(* Logix 5000 project; controller _GigaDiscovery vendor 1 type 14 code 244 rev 35.11; software revision 35.03; part 16 of 23 *)
(* tags used below, declared in another part *)
   E_Stop2_Test_Request : BOOL;
   E_Stop_Test_Request : BOOL;
   HMI_Pb_Platform_Open : BOOL;   // HMI Platform Open Command
   HMI_Platform_Close : BOOL;   // HMI Platform Close Command
   I_Compressor_Min_Pressure : BOOL;   // Line Pressure Switch - Minimum Pressure -S21504B
   I_Compressor_Work_Pressure : BOOL;   // Line Pressure Switch - Working Pressure -S21502B
   I_EStop_Pb_OCC1 : UDT_DCI_STOP_TEST;   // +OCC E-stop -S30301F
   I_EStop_Pb_OCC2 : UDT_DCI_STOP_TEST;   // +OCC2 E-Stop -S28502F
   I_HMI_Login_Enable : BOOL;   // Primary console Key selector Display Login -S30309F
   I_MCC_Temperature_OK : BOOL;   // MCC temeprature OK -S75003C
   I_OCC1_EntGate_PB : BOOL;   // OCC1 Entrance Gate Open/Close -S30701F
   I_OCC1_ExitGate_PB : BOOL;   // OCC1 ExitGate Open/Close -S30707F
   I_OCC1_Stop_Cycle_PB : BOOL;   // Stop Cycle -S30308F
   I_OCC2_ACONFIRM : BOOL;   // OCC2 Allow Main CONFIRM -S28602F
   I_OCC2_Disable : UDT_DCM;   // OCC 2 CONTROL DISABLE Page 310
   I_OCC2_RESTRAINTS_RELEASE : Sel_3_Pos_2_Input;   // -S28507F RESTRAINTS RELEASE UNLOCK -RUN- LOCK
   I_OCC2_Stop_Cycle_PB : BOOL;   // Stop Cycle -S28606F
   I_OCC_Aut_Man_Selector_Motion : UDT_DCM;   // S30801F
   I_OCC_Emergency_Brake : BOOL;   // I OCC Emergency Brake -S31207D
   I_OCC_LockOut_Motion : UDT_DCM;   // OCC -Lockout Motion -Q31203E
   I_OCC_Memory_Footpedal : BOOL;
   I_OCC_Operator_Enable_Key : BOOL;   // OCC Console Enabled -S30305F
   I_OCC_Temperature_OK : BOOL;   // OCC temperature OK -S31003E
   I_Operator_Footpedal : BOOL;   // Operator Footpedal -S30901F
   I_RESTRAINTS_MainValve_Cosed : BOOL;   // Main Valve Close Limit Switch -B40508I
   I_RESTRAINTS_PressureswitchCompressor : BOOL;   // RESTRAINTS Main Valve Pressure Switch -S40602J
   I_RESTRAINTS_Selector : Sel_3_Pos_2_Input;   // RESTRAINTS Selctor -S30505F Left = Open Right = Close Center = Nothing
   I_Start_PB : Start_AOI;   // Primary console Strat Push botton Right and Left -S30401F -S30403F
   MODE : BOOL;   // MODE 0 = AUTO 1 = MANUAL -S30801F
   No_Sfty : Std_to_Sfty;
   ONP : DINT;   // Optional Not Present
   Pb_Platform_Stop : BOOL;   // Platform Stop Command -S30608F
   Power_On_Delay : BOOL;
   Reset_Pulse : BOOL;
   RESTRAINTS_Rack : LapBar_Racks[41];
   RESTRAINTS_Sector : LapBars_Sector[9];
   Start_Stop_Cycle : Sequencer;
   ToBe_Define_Sfty : DINT[10];

PROGRAM S_Input   (* main routine Main, safety *)
VAR
   E_Stop_Secondary_Released : BOOL := 1;
   Home_Timer : TIMER := (PRE := 10000, ACC := 10000, EN := 1, DN := 1);
   Os : DINT := 14;
   Reset_Start_AOI : BOOL;   // Start AOI Instruction Reset
   Reset_Status : TIMER := (PRE := 1500, ACC := 1520);
   timer : TIMER[10] := ([0].PRE := 30000, [0].ACC := 30000, [0].EN := 1, [0].DN := 1, [1].PRE := 8000, [1].ACC := 8000, [1].EN := 1, [1].DN := 1, [2].PRE := 3000, [2].EN := 1, [2].DN := 1, [3].PRE := 4000, [4].PRE := 2000, [5].PRE := 5000, [6].PRE := 500, [7].PRE := 500, [8].PRE := 1600);
   Timer2 : TIMER := (PRE := 5000, ACC := 5000, EN := 1, DN := 1);
END_VAR

ROUTINE _01_OCC   (* ladder *)
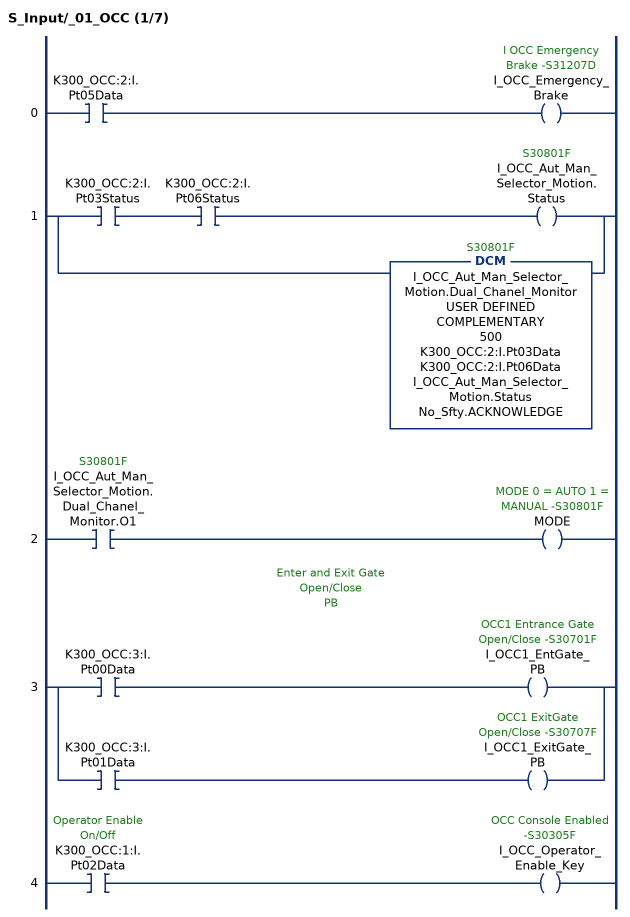
   0: XIC(K300_OCC:2:I.Pt05Data)OTE(I_OCC_Emergency_Brake);
   1: [XIC(K300_OCC:2:I.Pt03Status) XIC(K300_OCC:2:I.Pt06Status) OTE(I_OCC_Aut_Man_Selector_Motion.Status) ,DCM(I_OCC_Aut_Man_Selector_Motion.Dual_Chanel_Monitor,USER DEFINED,COMPLEMENTARY,500,K300_OCC:2:I.Pt03Data,K300_OCC:2:I.Pt06Data,I_OCC_Aut_Man_Selector_Motion.Status,No_Sfty.ACKNOWLEDGE) ];
   2: XIC(I_OCC_Aut_Man_Selector_Motion.Dual_Chanel_Monitor.O1)OTE(MODE);
   // Enter and Exit Gate
   // Open/Close
   // PB
   3: [XIC(K300_OCC:3:I.Pt00Data) OTE(I_OCC1_EntGate_PB) ,XIC(K300_OCC:3:I.Pt01Data) OTE(I_OCC1_ExitGate_PB) ];
   4: XIC(K300_OCC:1:I.Pt02Data)OTE(I_OCC_Operator_Enable_Key);
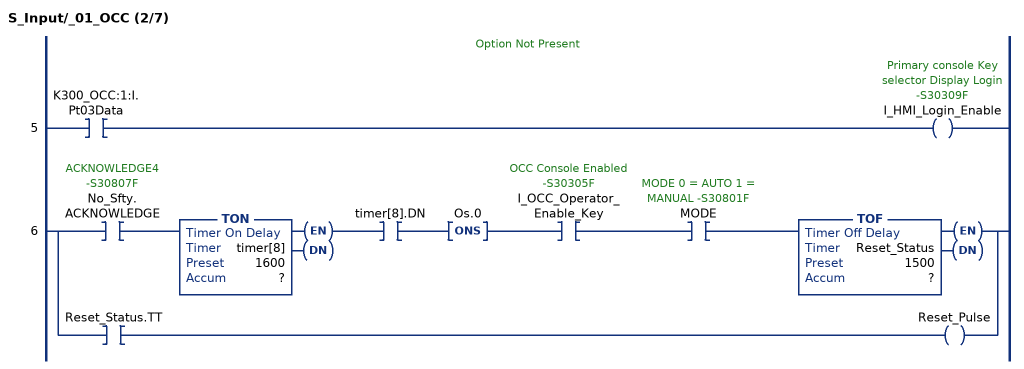
   // Option Not Present
   5: XIC(K300_OCC:1:I.Pt03Data)OTE(I_HMI_Login_Enable);
   6: [XIC(No_Sfty.ACKNOWLEDGE) TON(timer[8],?,?) XIC(timer[8].DN) ONS(Os.0) XIC(I_OCC_Operator_Enable_Key) XIC(MODE) TOF(Reset_Status,?,?) ,XIC(Reset_Status.TT) OTE(Reset_Pulse) ];
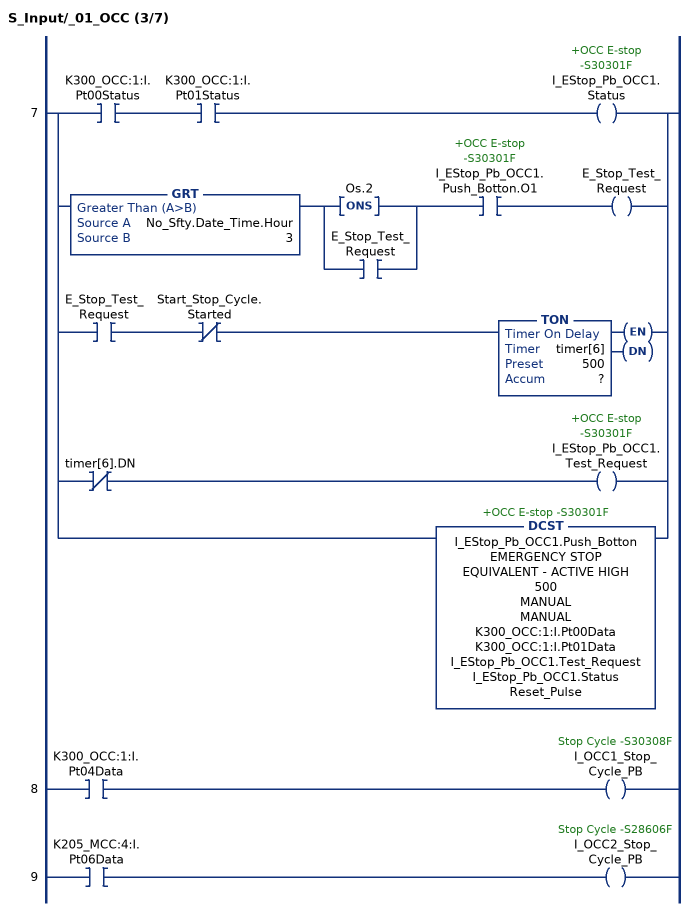
   7: [XIC(K300_OCC:1:I.Pt00Status) XIC(K300_OCC:1:I.Pt01Status) OTE(I_EStop_Pb_OCC1.Status) ,GRT(No_Sfty.Date_Time.Hour,3) [ONS(Os.2) ,XIC(E_Stop_Test_Request) ] XIC(I_EStop_Pb_OCC1.Push_Botton.O1) OTE(E_Stop_Test_Request) ,XIC(E_Stop_Test_Request) XIO(Start_Stop_Cycle.Started) TON(timer[6],?,?) ,XIO(timer[6].DN) OTE(I_EStop_Pb_OCC1.Test_Request) ,DCST(I_EStop_Pb_OCC1.Push_Botton,EMERGENCY STOP,EQUIVALENT - ACTIVE HIGH,500,MANUAL,MANUAL,K300_OCC:1:I.Pt00Data,K300_OCC:1:I.Pt01Data,I_EStop_Pb_OCC1.Test_Request,I_EStop_Pb_OCC1.Status,Reset_Pulse) ];
   8: XIC(K300_OCC:1:I.Pt04Data)OTE(I_OCC1_Stop_Cycle_PB);
   9: XIC(K205_MCC:4:I.Pt06Data)OTE(I_OCC2_Stop_Cycle_PB);
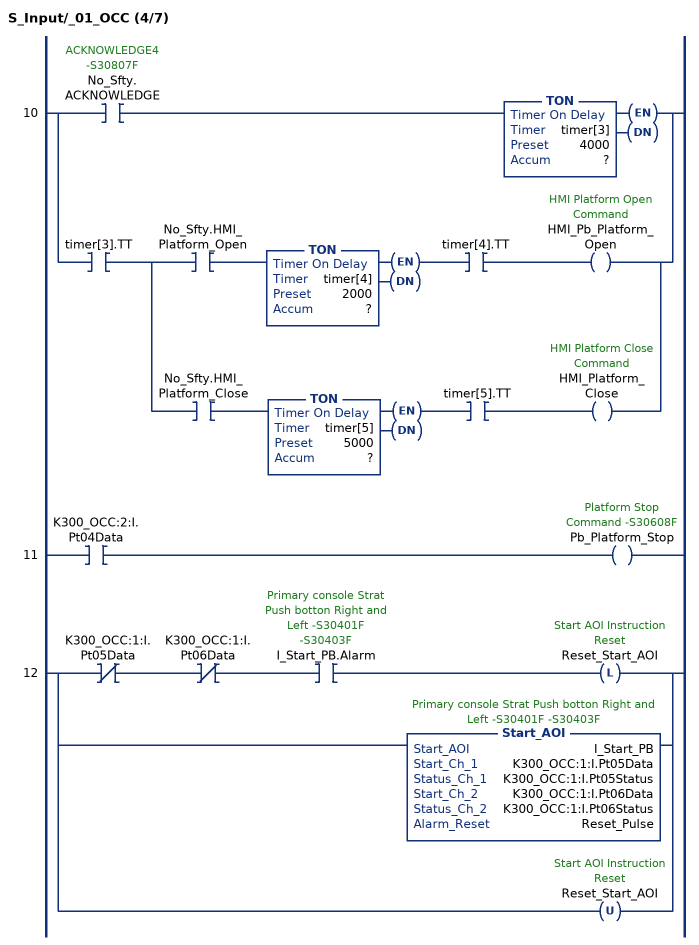
   10: [XIC(No_Sfty.ACKNOWLEDGE) TON(timer[3],?,?) ,XIC(timer[3].TT) [XIC(No_Sfty.HMI_Platform_Open) TON(timer[4],?,?) XIC(timer[4].TT) OTE(HMI_Pb_Platform_Open) ,XIC(No_Sfty.HMI_Platform_Close) TON(timer[5],?,?) XIC(timer[5].TT) OTE(HMI_Platform_Close) ] ];
   11: XIC(K300_OCC:2:I.Pt04Data)OTE(Pb_Platform_Stop);
   12: [XIO(K300_OCC:1:I.Pt05Data) XIO(K300_OCC:1:I.Pt06Data) XIC(I_Start_PB.Alarm) OTL(Reset_Start_AOI) ,Start_AOI(I_Start_PB,K300_OCC:1:I.Pt05Data,K300_OCC:1:I.Pt05Status,K300_OCC:1:I.Pt06Data,K300_OCC:1:I.Pt06Status,Reset_Pulse) ,OTU(Reset_Start_AOI) ];
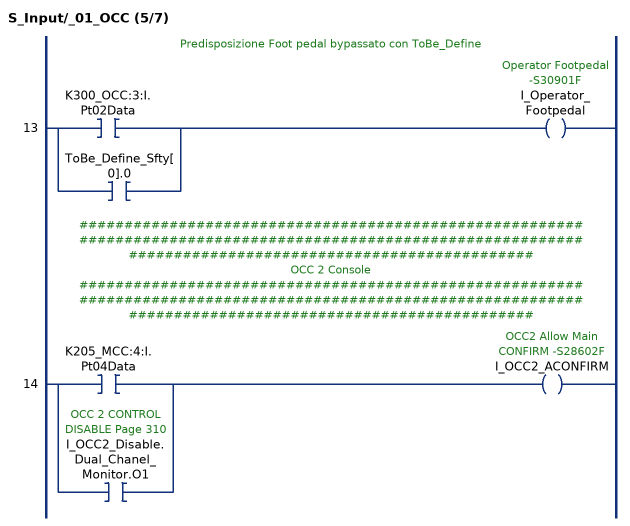
   // Predisposizione Foot pedal bypassato con ToBe_Define
   13: [XIC(K300_OCC:3:I.Pt02Data) ,XIC(ToBe_Define_Sfty[0].0) ]OTE(I_Operator_Footpedal);
   // #############################################################################################################################################################
   // OCC 2 Console
   // #############################################################################################################################################################
   14: [XIC(K205_MCC:4:I.Pt04Data) ,XIC(I_OCC2_Disable.Dual_Chanel_Monitor.O1) ]OTE(I_OCC2_ACONFIRM);
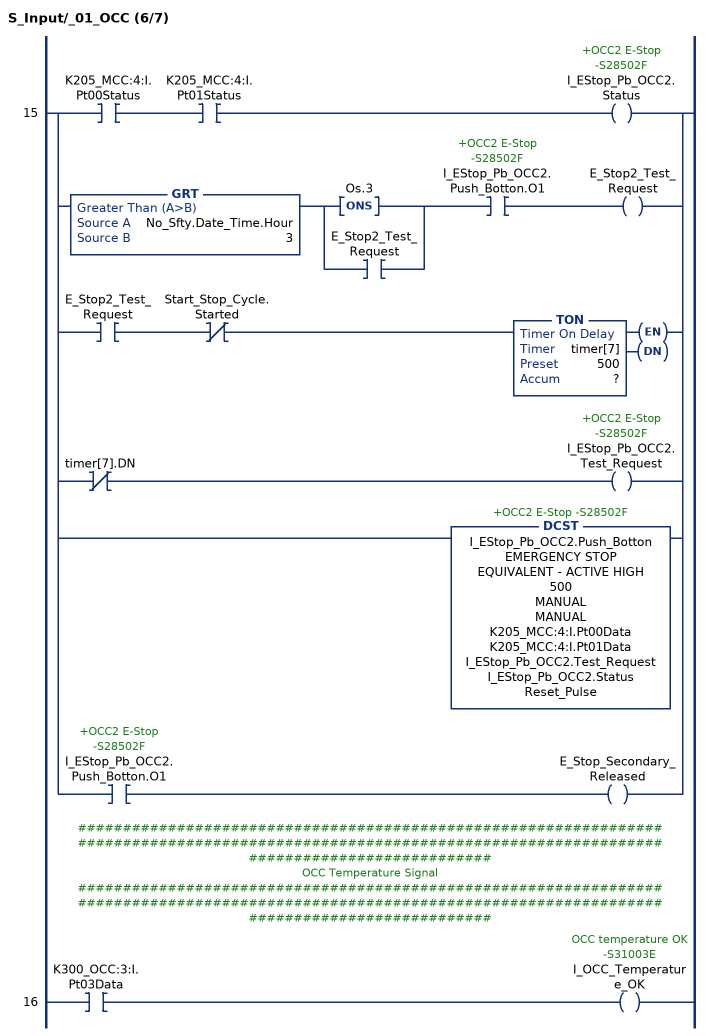
   15: [XIC(K205_MCC:4:I.Pt00Status) XIC(K205_MCC:4:I.Pt01Status) OTE(I_EStop_Pb_OCC2.Status) ,GRT(No_Sfty.Date_Time.Hour,3) [ONS(Os.3) ,XIC(E_Stop2_Test_Request) ] XIC(I_EStop_Pb_OCC2.Push_Botton.O1) OTE(E_Stop2_Test_Request) ,XIC(E_Stop2_Test_Request) XIO(Start_Stop_Cycle.Started) TON(timer[7],?,?) ,XIO(timer[7].DN) OTE(I_EStop_Pb_OCC2.Test_Request) ,DCST(I_EStop_Pb_OCC2.Push_Botton,EMERGENCY STOP,EQUIVALENT - ACTIVE HIGH,500,MANUAL,MANUAL,K205_MCC:4:I.Pt00Data,K205_MCC:4:I.Pt01Data,I_EStop_Pb_OCC2.Test_Request,I_EStop_Pb_OCC2.Status,Reset_Pulse) ,XIC(I_EStop_Pb_OCC2.Push_Botton.O1) OTE(E_Stop_Secondary_Released) ];
   // #############################################################################################################################################################
   // OCC Temperature Signal
   // #############################################################################################################################################################
   16: XIC(K300_OCC:3:I.Pt03Data)OTE(I_OCC_Temperature_OK);
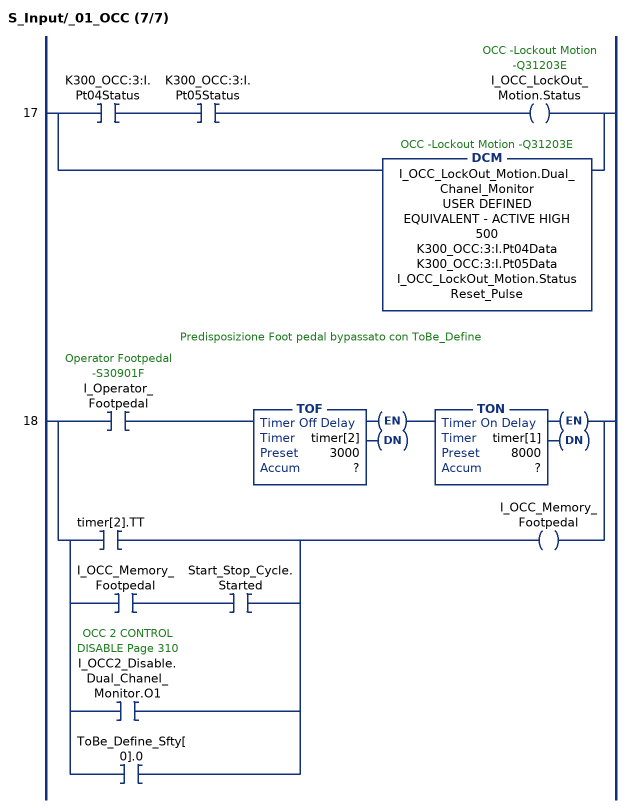
   17: [XIC(K300_OCC:3:I.Pt04Status) XIC(K300_OCC:3:I.Pt05Status) OTE(I_OCC_LockOut_Motion.Status) ,DCM(I_OCC_LockOut_Motion.Dual_Chanel_Monitor,USER DEFINED,EQUIVALENT - ACTIVE HIGH,500,K300_OCC:3:I.Pt04Data,K300_OCC:3:I.Pt05Data,I_OCC_LockOut_Motion.Status,Reset_Pulse) ];
   // Predisposizione Foot pedal bypassato con ToBe_Define
   18: [XIC(I_Operator_Footpedal) TOF(timer[2],?,?) TON(timer[1],?,?) ,[XIC(timer[2].TT) ,XIC(I_OCC_Memory_Footpedal) XIC(Start_Stop_Cycle.Started) ,XIC(I_OCC2_Disable.Dual_Chanel_Monitor.O1) ,XIC(ToBe_Define_Sfty[0].0) ] OTE(I_OCC_Memory_Footpedal) ];
END_ROUTINE

ROUTINE _02_MCC   (* ladder *)
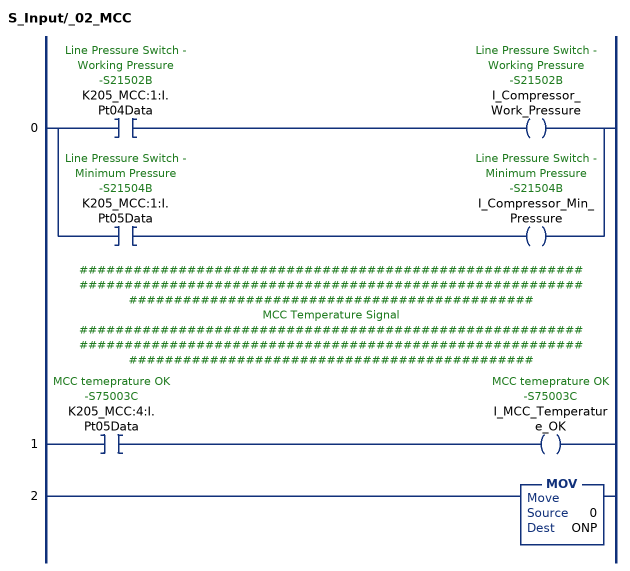
   0: [XIC(K205_MCC:1:I.Pt04Data) OTE(I_Compressor_Work_Pressure) ,XIC(K205_MCC:1:I.Pt05Data) OTE(I_Compressor_Min_Pressure) ];
   // #############################################################################################################################################################
   // MCC Temperature Signal
   // #############################################################################################################################################################
   1: XIC(K205_MCC:4:I.Pt05Data)OTE(I_MCC_Temperature_OK);
   2: MOV(0,ONP);
END_ROUTINE

ROUTINE _03_RESTRAINT_RELEASE   (* ladder *)
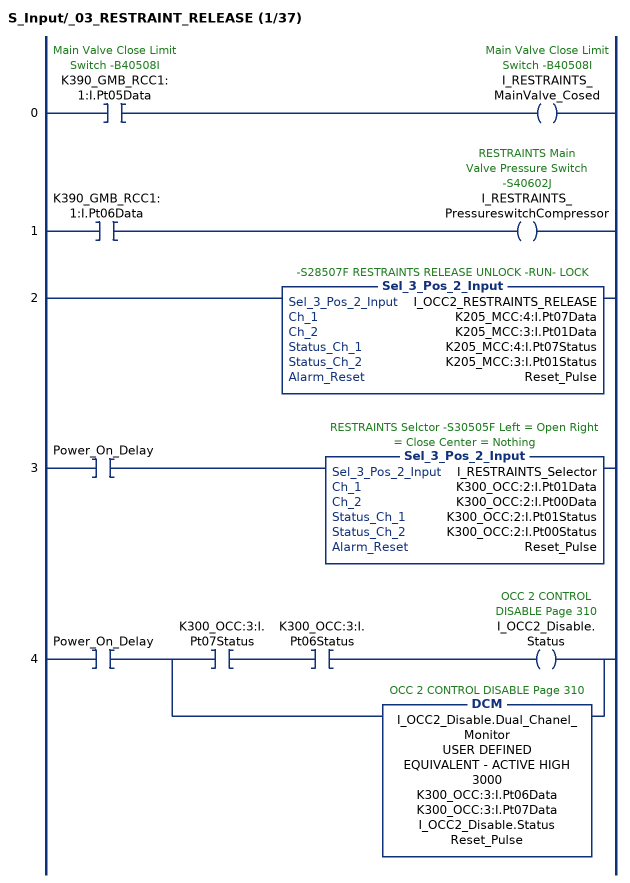
   0: XIC(K390_GMB_RCC1:1:I.Pt05Data)OTE(I_RESTRAINTS_MainValve_Cosed);
   1: XIC(K390_GMB_RCC1:1:I.Pt06Data)OTE(I_RESTRAINTS_PressureswitchCompressor);
   2: Sel_3_Pos_2_Input(I_OCC2_RESTRAINTS_RELEASE,K205_MCC:4:I.Pt07Data,K205_MCC:3:I.Pt01Data,K205_MCC:4:I.Pt07Status,K205_MCC:3:I.Pt01Status,Reset_Pulse);
   3: XIC(Power_On_Delay)Sel_3_Pos_2_Input(I_RESTRAINTS_Selector,K300_OCC:2:I.Pt01Data,K300_OCC:2:I.Pt00Data,K300_OCC:2:I.Pt01Status,K300_OCC:2:I.Pt00Status,Reset_Pulse);
   4: XIC(Power_On_Delay)[XIC(K300_OCC:3:I.Pt07Status) XIC(K300_OCC:3:I.Pt06Status) OTE(I_OCC2_Disable.Status) ,DCM(I_OCC2_Disable.Dual_Chanel_Monitor,USER DEFINED,EQUIVALENT - ACTIVE HIGH,3000,K300_OCC:3:I.Pt06Data,K300_OCC:3:I.Pt07Data,I_OCC2_Disable.Status,Reset_Pulse) ];
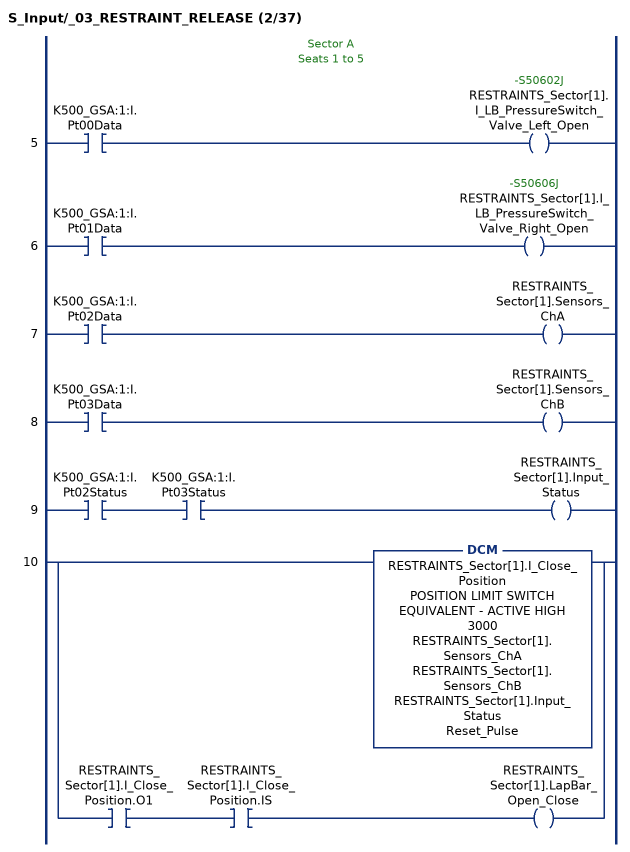
   // Sector A
   // Seats 1 to 5
   5: XIC(K500_GSA:1:I.Pt00Data)OTE(RESTRAINTS_Sector[1].I_LB_PressureSwitch_Valve_Left_Open);
   6: XIC(K500_GSA:1:I.Pt01Data)OTE(RESTRAINTS_Sector[1].I_LB_PressureSwitch_Valve_Right_Open);
   7: XIC(K500_GSA:1:I.Pt02Data)OTE(RESTRAINTS_Sector[1].Sensors_ChA);
   8: XIC(K500_GSA:1:I.Pt03Data)OTE(RESTRAINTS_Sector[1].Sensors_ChB);
   9: XIC(K500_GSA:1:I.Pt02Status)XIC(K500_GSA:1:I.Pt03Status)OTE(RESTRAINTS_Sector[1].Input_Status);
   10: [DCM(RESTRAINTS_Sector[1].I_Close_Position,POSITION LIMIT SWITCH,EQUIVALENT - ACTIVE HIGH,3000,RESTRAINTS_Sector[1].Sensors_ChA,RESTRAINTS_Sector[1].Sensors_ChB,RESTRAINTS_Sector[1].Input_Status,Reset_Pulse) ,XIC(RESTRAINTS_Sector[1].I_Close_Position.O1) XIC(RESTRAINTS_Sector[1].I_Close_Position.IS) OTE(RESTRAINTS_Sector[1].LapBar_Open_Close) ];
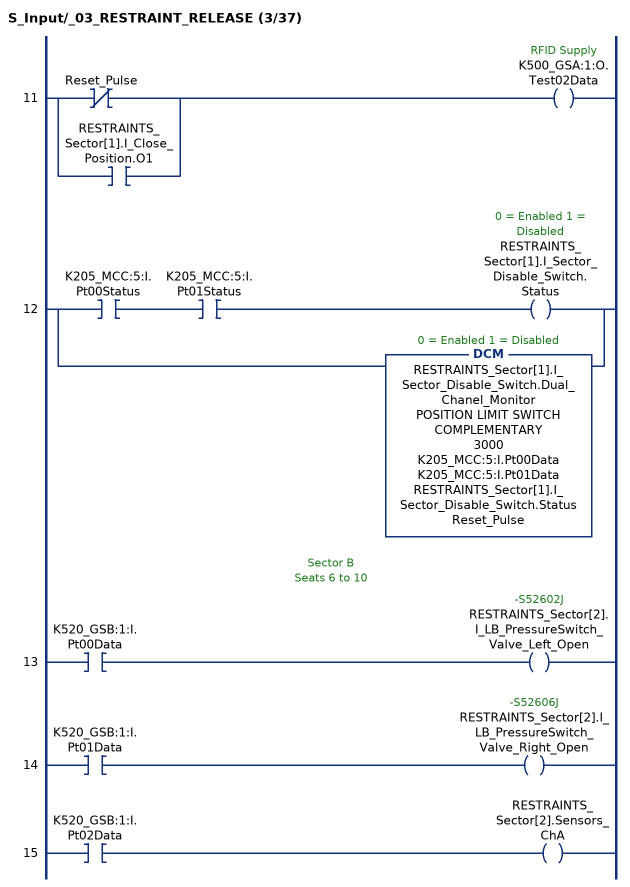
   11: [XIO(Reset_Pulse) ,XIC(RESTRAINTS_Sector[1].I_Close_Position.O1) ]OTE(K500_GSA:1:O.Test02Data);
   12: [XIC(K205_MCC:5:I.Pt00Status) XIC(K205_MCC:5:I.Pt01Status) OTE(RESTRAINTS_Sector[1].I_Sector_Disable_Switch.Status) ,DCM(RESTRAINTS_Sector[1].I_Sector_Disable_Switch.Dual_Chanel_Monitor,POSITION LIMIT SWITCH,COMPLEMENTARY,3000,K205_MCC:5:I.Pt00Data,K205_MCC:5:I.Pt01Data,RESTRAINTS_Sector[1].I_Sector_Disable_Switch.Status,Reset_Pulse) ];
   // Sector B
   // Seats 6 to 10
   13: XIC(K520_GSB:1:I.Pt00Data)OTE(RESTRAINTS_Sector[2].I_LB_PressureSwitch_Valve_Left_Open);
   14: XIC(K520_GSB:1:I.Pt01Data)OTE(RESTRAINTS_Sector[2].I_LB_PressureSwitch_Valve_Right_Open);
   15: XIC(K520_GSB:1:I.Pt02Data)OTE(RESTRAINTS_Sector[2].Sensors_ChA);
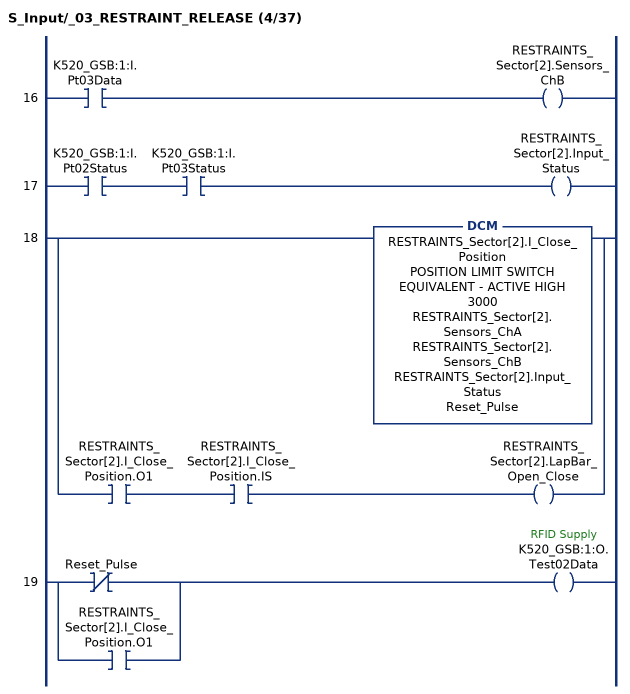
   16: XIC(K520_GSB:1:I.Pt03Data)OTE(RESTRAINTS_Sector[2].Sensors_ChB);
   17: XIC(K520_GSB:1:I.Pt02Status)XIC(K520_GSB:1:I.Pt03Status)OTE(RESTRAINTS_Sector[2].Input_Status);
   18: [DCM(RESTRAINTS_Sector[2].I_Close_Position,POSITION LIMIT SWITCH,EQUIVALENT - ACTIVE HIGH,3000,RESTRAINTS_Sector[2].Sensors_ChA,RESTRAINTS_Sector[2].Sensors_ChB,RESTRAINTS_Sector[2].Input_Status,Reset_Pulse) ,XIC(RESTRAINTS_Sector[2].I_Close_Position.O1) XIC(RESTRAINTS_Sector[2].I_Close_Position.IS) OTE(RESTRAINTS_Sector[2].LapBar_Open_Close) ];
   19: [XIO(Reset_Pulse) ,XIC(RESTRAINTS_Sector[2].I_Close_Position.O1) ]OTE(K520_GSB:1:O.Test02Data);